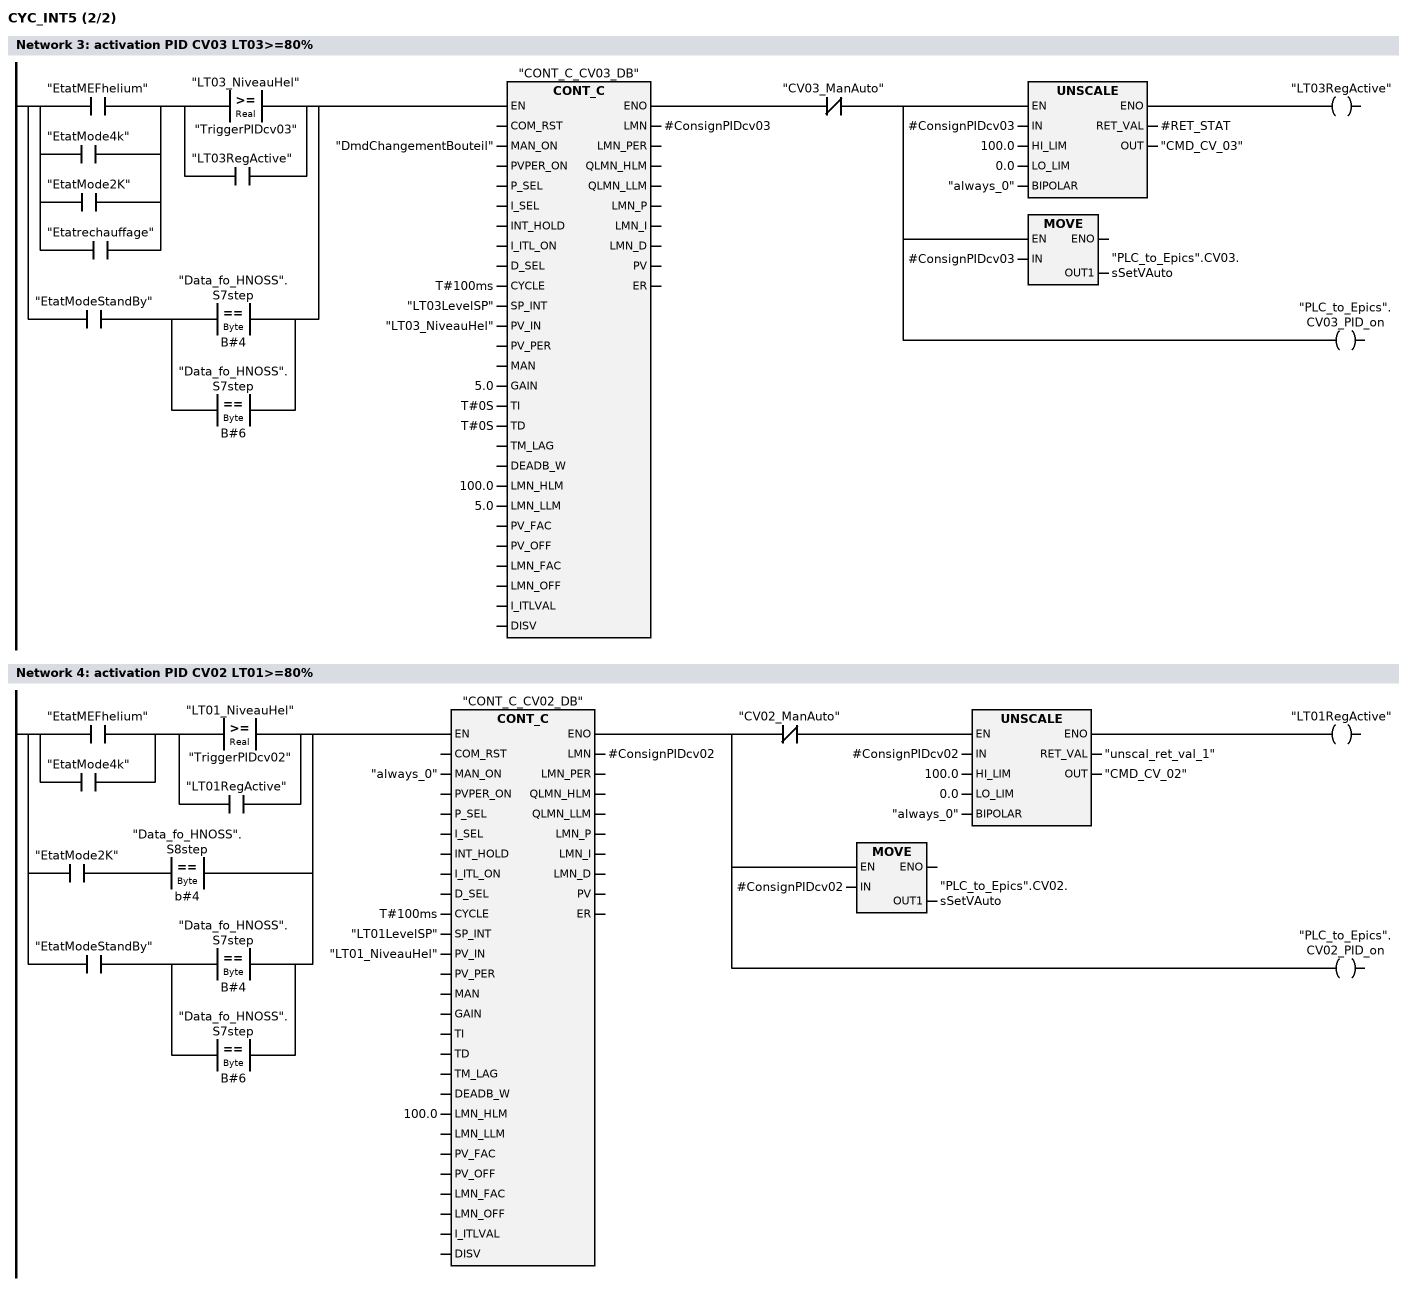
   // ENO of a box is taken as its EN; it also drops when the box reports an error
   #_w1 := (("EtatMEFhelium" OR "EtatMode4k" OR "EtatMode2K" OR "Etatrechauffage") AND (("LT03_NiveauHel" >= "TriggerPIDcv03") OR "LT03RegActive")) OR ("EtatModeStandBy" AND (("Data_fo_HNOSS".S7step = B#4) OR ("Data_fo_HNOSS".S7step = B#6)));
   IF #_w1 THEN
       "CONT_C_CV03_DB"(MAN_ON := "DmdChangementBouteil",   // CONT_C
                        CYCLE := T#100ms,
                        SP_INT := "LT03LevelSP",
                        PV_IN := "LT03_NiveauHel",
                        GAIN := 5.0,
                        TI := T#0S,
                        TD := T#0S,
                        LMN_HLM := 100.0,
                        LMN_LLM := 5.0,
                        LMN => #ConsignPIDcv03);
   END_IF;
   #_w2 := #_w1 AND NOT "CV03_ManAuto";
   IF #_w2 THEN
       #RET_STAT := UNSCALE(IN := #ConsignPIDcv03,
                            HI_LIM := 100.0,
                            LO_LIM := 0.0,
                            BIPOLAR := "always_0",
                            OUT => "CMD_CV_03");
   END_IF;
   "LT03RegActive" := #_w2;
   IF #_w2 THEN "PLC_to_Epics".CV03.sSetVAuto := #ConsignPIDcv03; END_IF;
   "PLC_to_Epics".CV03_PID_on := #_w2;
END_REGION

REGION Network 4: activation PID CV02 LT01>=80%
   // ENO of a box is taken as its EN; it also drops when the box reports an error
   #_w1 := (("EtatMEFhelium" OR "EtatMode4k") AND (("LT01_NiveauHel" >= "TriggerPIDcv02") OR "LT01RegActive")) OR ("EtatMode2K" AND ("Data_fo_HNOSS".S8step = b#4)) OR ("EtatModeStandBy" AND (("Data_fo_HNOSS".S7step = B#4) OR ("Data_fo_HNOSS".S7step = B#6)));
   IF #_w1 THEN
       "CONT_C_CV02_DB"(MAN_ON := "always_0",   // CONT_C
                        CYCLE := T#100ms,
                        SP_INT := "LT01LevelSP",
                        PV_IN := "LT01_NiveauHel",
                        LMN_HLM := 100.0,
                        LMN => #ConsignPIDcv02);
   END_IF;
   #_w2 := #_w1 AND NOT "CV02_ManAuto";
   IF #_w2 THEN
       "unscal_ret_val_1" := UNSCALE(IN := #ConsignPIDcv02,
                               HI_LIM := 100.0,
                               LO_LIM := 0.0,
                               BIPOLAR := "always_0",
                               OUT => "CMD_CV_02");
   END_IF;
   "LT01RegActive" := #_w2;
   IF #_w1 THEN "PLC_to_Epics".CV02.sSetVAuto := #ConsignPIDcv02; END_IF;
   "PLC_to_Epics".CV02_PID_on := #_w1;
END_REGION
END_ORGANIZATION_BLOCK

ORGANIZATION_BLOCK "HW_INT0"   // OB40, LAD
TITLE = "Hardware Interrupt"
{ S7_Optimized_Access := 'FALSE' }
VERSION : 0.1
BEGIN
END_ORGANIZATION_BLOCK

ORGANIZATION_BLOCK "I/O_FLT1"   // OB82, LAD
TITLE = "I/O Point Fault"
{ S7_Optimized_Access := 'FALSE' }
VERSION : 0.1
BEGIN

REGION Network 1 (STL): Appeler le bloc de diagnostic système / Call system diagnostics block
         CALL  "RSE_FB", "RSE_DB";
END_REGION
END_ORGANIZATION_BLOCK

ORGANIZATION_BLOCK "OBNL_FLT"   // OB85, LAD
TITLE = "Organization Block (OB) Not Loaded Fault"
{ S7_Optimized_Access := 'FALSE' }
VERSION : 0.1
BEGIN
END_ORGANIZATION_BLOCK

ORGANIZATION_BLOCK "RACK_FLT"   // OB86, LAD
TITLE = "Loss Of Rack Fault"
{ S7_Optimized_Access := 'FALSE' }
VERSION : 0.1
BEGIN

REGION Network 1 (STL): Appeler le bloc de diagnostic système / Call system diagnostics block
         CALL  "RSE_FB", "RSE_DB";
END_REGION
END_ORGANIZATION_BLOCK

ORGANIZATION_BLOCK "COMPLETE RESTART"   // OB100, STL
TITLE = "Complete Restart"
{ S7_Optimized_Access := 'FALSE' }
VERSION : 0.1
BEGIN

REGION Network 1
         SET;
         S     "INIT";
END_REGION
END_ORGANIZATION_BLOCK

(* ===== HMI "HMI_RT_1" =====

graphic list "Vanne horizontale maxi_0": 1 'Vanne horizontale verte_2'; 0 'Vanne horizontale rouge_2'; 2 'Vanne horizontale rouge_2'; 3 'Vanne horizontale verte_2'; 4 'Vanne horizontale grise_2'; 5 'Vanne horizontale grise_2'

ScreenModuleEditorView "Bloc Vanne horizontale" 1024x768
   GraphicIOField "Modèle_Champ E/S graphique_13" at 10,10 size 50x35
*)

(* ===== HMI "HMI_RT_1" =====

graphic list "Vanne verticale maxi_0": 1 'Vanne verticale verte_1'; 2 'Vanne verticale rouge_1'; 0 'Vanne verticale rouge_1'; 3 'Vanne verticale verte_1'; 4 'Vanne verticale grise_1'; 5 'Vanne verticale grise_1'

ScreenModuleEditorView "Bloc Vanne verticale" 1024x768
   GraphicIOField "Champ E/S graphique_10" at 10,10 size 35x50
*)